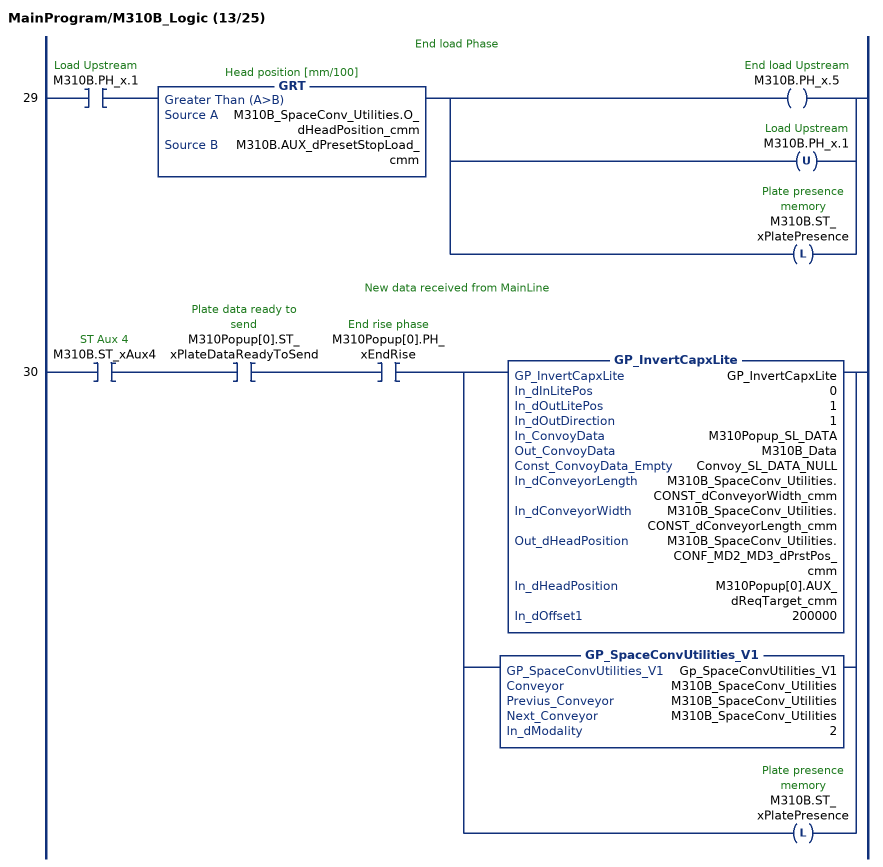
   // End load Phase
   29: XIC(M310B.PH_x.1)GRT(M310B_SpaceConv_Utilities.O_dHeadPosition_cmm,M310B.AUX_dPresetStopLoad_cmm)[OTE(M310B.PH_x.5) ,OTU(M310B.PH_x.1) ,OTL(M310B.ST_xPlatePresence) ];
   // New data received from MainLine
   30: XIC(M310B.ST_xAux4)XIC(M310Popup[0].ST_xPlateDataReadyToSend)XIC(M310Popup[0].PH_xEndRise)[GP_InvertCapxLite(GP_InvertCapxLite,0,1,1,M310Popup_SL_DATA,M310B_Data,Convoy_SL_DATA_NULL,M310B_SpaceConv_Utilities.CONST_dConveyorWidth_cmm,M310B_SpaceConv_Utilities.CONST_dConveyorLength_cmm,M310B_SpaceConv_Utilities.CONF_MD2_MD3_dPrstPos_cmm,M310Popup[0].AUX_dReqTarget_cmm,200000) ,GP_SpaceConvUtilities_V1(Gp_SpaceConvUtilities_V1,M310B_SpaceConv_Utilities,M310B_SpaceConv_Utilities,M310B_SpaceConv_Utilities,2) ,OTL(M310B.ST_xPlatePresence) ];
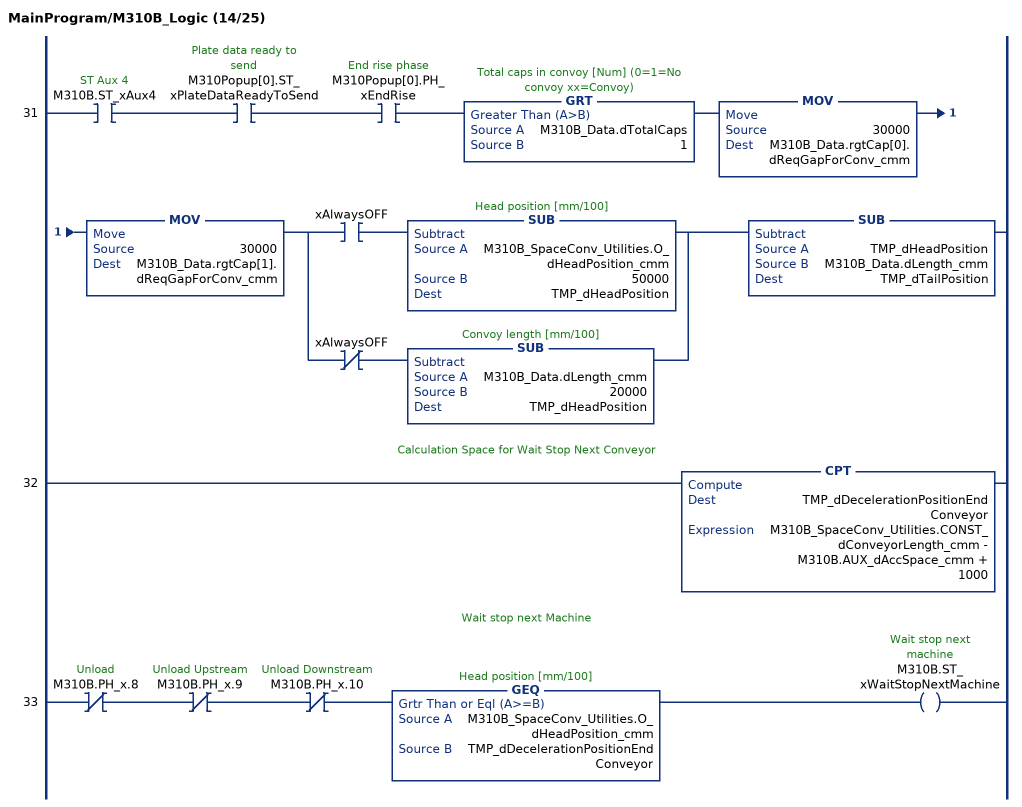
   31: XIC(M310B.ST_xAux4)XIC(M310Popup[0].ST_xPlateDataReadyToSend)XIC(M310Popup[0].PH_xEndRise)GRT(M310B_Data.dTotalCaps,1)MOV(30000,M310B_Data.rgtCap[0].dReqGapForConv_cmm)MOV(30000,M310B_Data.rgtCap[1].dReqGapForConv_cmm)[XIC(xAlwaysOFF) SUB(M310B_SpaceConv_Utilities.O_dHeadPosition_cmm,50000,TMP_dHeadPosition) ,XIO(xAlwaysOFF) SUB(M310B_Data.dLength_cmm,20000,TMP_dHeadPosition) ]SUB(TMP_dHeadPosition,M310B_Data.dLength_cmm,TMP_dTailPosition);
   // Calculation Space for Wait Stop Next Conveyor
   32: CPT(TMP_dDecelerationPositionEndConveyor,M310B_SpaceConv_Utilities.CONST_dConveyorLength_cmm - M310B.AUX_dAccSpace_cmm + 1000);
   // Wait stop next Machine
   33: XIO(M310B.PH_x.8)XIO(M310B.PH_x.9)XIO(M310B.PH_x.10)GEQ(M310B_SpaceConv_Utilities.O_dHeadPosition_cmm,TMP_dDecelerationPositionEndConveyor)OTE(M310B.ST_xWaitStopNextMachine);
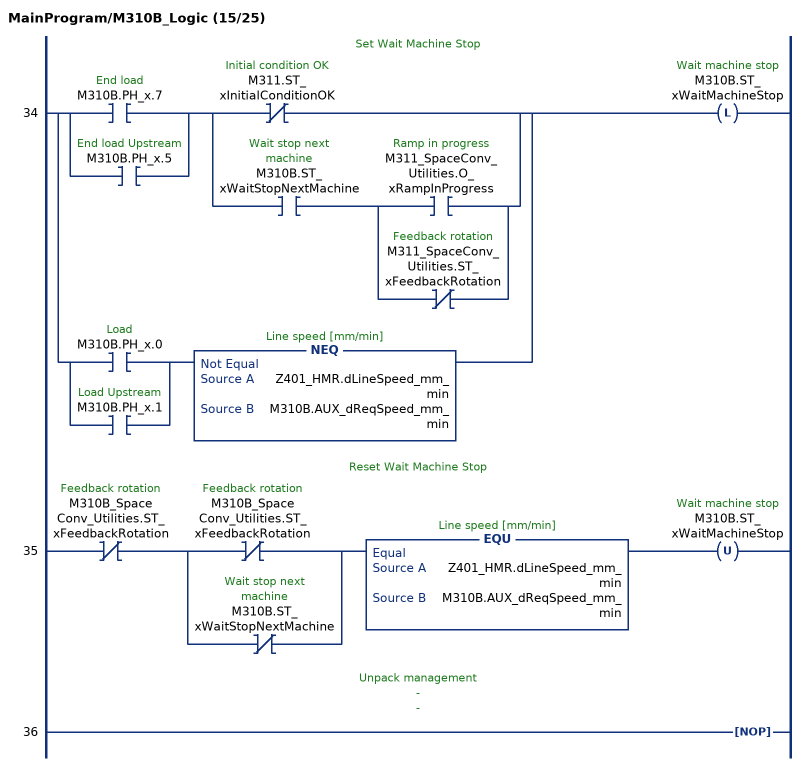
   // Set Wait Machine Stop
   34: [[XIC(M310B.PH_x.7) ,XIC(M310B.PH_x.5) ] [XIO(M311.ST_xInitialConditionOK) ,XIC(M310B.ST_xWaitStopNextMachine) [XIC(M311_SpaceConv_Utilities.O_xRampInProgress) ,XIO(M311_SpaceConv_Utilities.ST_xFeedbackRotation) ] ] ,[XIC(M310B.PH_x.0) ,XIC(M310B.PH_x.1) ] NEQ(Z401_HMR.dLineSpeed_mm_min,M310B.AUX_dReqSpeed_mm_min) ]OTL(M310B.ST_xWaitMachineStop);
   // Reset Wait Machine Stop
   35: XIO(M310B_SpaceConv_Utilities.ST_xFeedbackRotation)[XIO(M310B_SpaceConv_Utilities.ST_xFeedbackRotation) ,XIO(M310B.ST_xWaitStopNextMachine) ]EQU(Z401_HMR.dLineSpeed_mm_min,M310B.AUX_dReqSpeed_mm_min)OTU(M310B.ST_xWaitMachineStop);
   // Unpack management
   // -
   // -
   36: NOP();
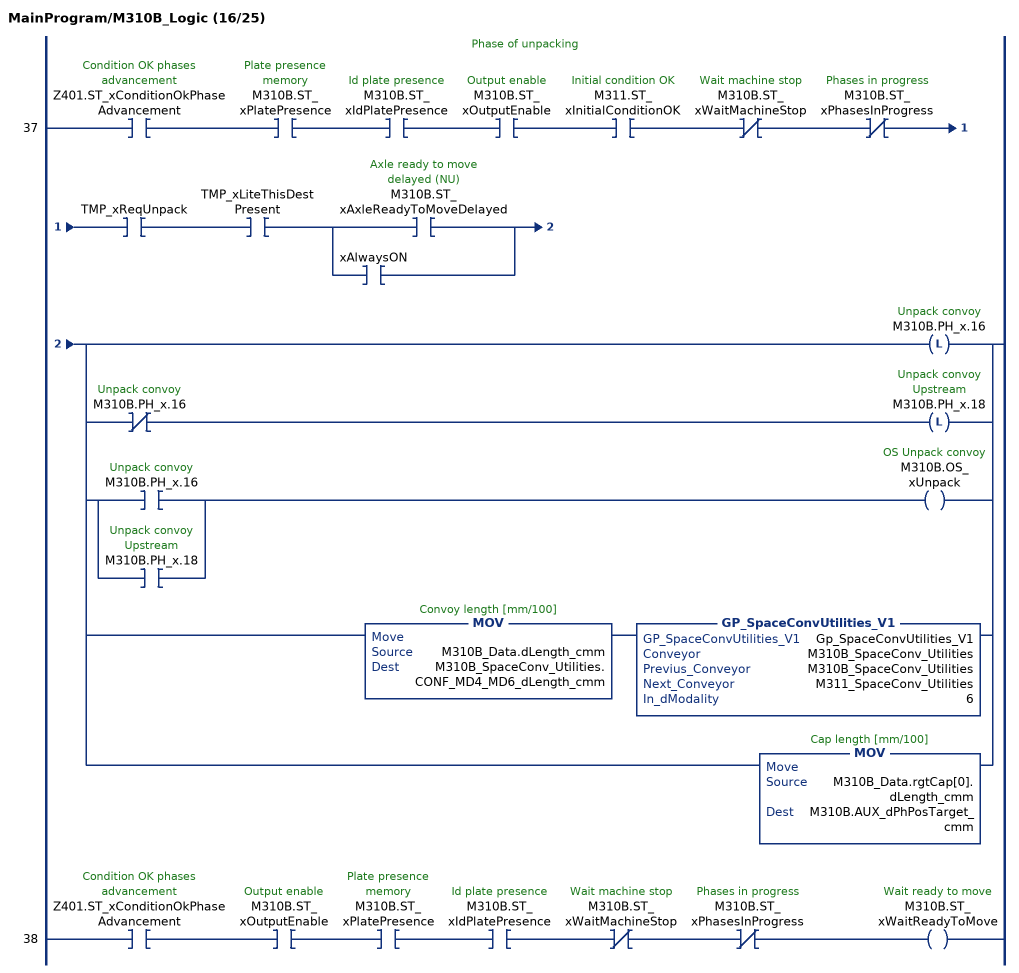
   // Phase of unpacking
   37: XIC(Z401.ST_xConditionOkPhaseAdvancement)XIC(M310B.ST_xPlatePresence)XIC(M310B.ST_xIdPlatePresence)XIC(M310B.ST_xOutputEnable)XIC(M311.ST_xInitialConditionOK)XIO(M310B.ST_xWaitMachineStop)XIO(M310B.ST_xPhasesInProgress)XIC(TMP_xReqUnpack)XIC(TMP_xLiteThisDestPresent)[XIC(M310B.ST_xAxleReadyToMoveDelayed) ,XIC(xAlwaysON) ][OTL(M310B.PH_x.16) ,XIO(M310B.PH_x.16) OTL(M310B.PH_x.18) ,[XIC(M310B.PH_x.16) ,XIC(M310B.PH_x.18) ] OTE(M310B.OS_xUnpack) ,MOV(M310B_Data.dLength_cmm,M310B_SpaceConv_Utilities.CONF_MD4_MD6_dLength_cmm) GP_SpaceConvUtilities_V1(Gp_SpaceConvUtilities_V1,M310B_SpaceConv_Utilities,M310B_SpaceConv_Utilities,M311_SpaceConv_Utilities,6) ,MOV(M310B_Data.rgtCap[0].dLength_cmm,M310B.AUX_dPhPosTarget_cmm) ];
   38: XIC(Z401.ST_xConditionOkPhaseAdvancement)XIC(M310B.ST_xOutputEnable)XIC(M310B.ST_xPlatePresence)XIC(M310B.ST_xIdPlatePresence)XIO(M310B.ST_xWaitMachineStop)XIO(M310B.ST_xPhasesInProgress)OTE(M310B.ST_xWaitReadyToMove);
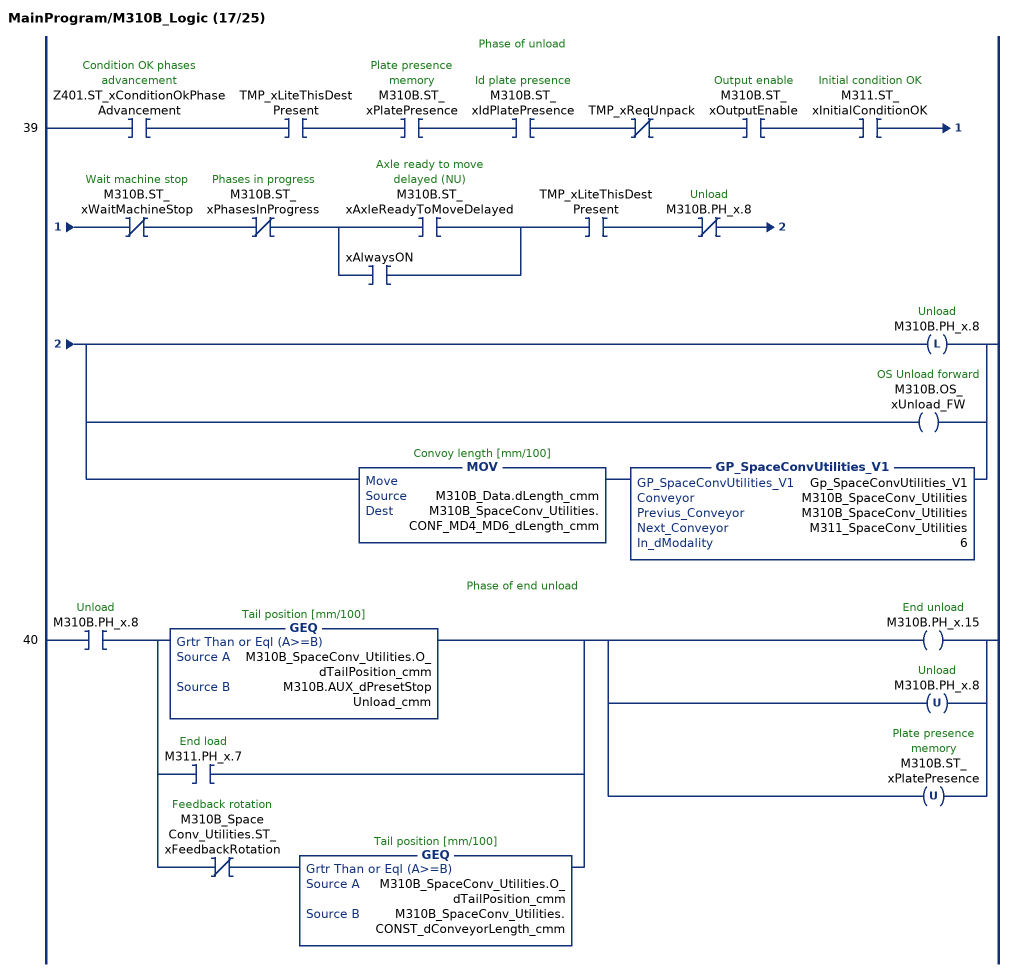
   // Phase of unload
   39: XIC(Z401.ST_xConditionOkPhaseAdvancement)XIC(TMP_xLiteThisDestPresent)XIC(M310B.ST_xPlatePresence)XIC(M310B.ST_xIdPlatePresence)XIO(TMP_xReqUnpack)XIC(M310B.ST_xOutputEnable)XIC(M311.ST_xInitialConditionOK)XIO(M310B.ST_xWaitMachineStop)XIO(M310B.ST_xPhasesInProgress)[XIC(M310B.ST_xAxleReadyToMoveDelayed) ,XIC(xAlwaysON) ]XIC(TMP_xLiteThisDestPresent)XIO(M310B.PH_x.8)[OTL(M310B.PH_x.8) ,OTE(M310B.OS_xUnload_FW) ,MOV(M310B_Data.dLength_cmm,M310B_SpaceConv_Utilities.CONF_MD4_MD6_dLength_cmm) GP_SpaceConvUtilities_V1(Gp_SpaceConvUtilities_V1,M310B_SpaceConv_Utilities,M310B_SpaceConv_Utilities,M311_SpaceConv_Utilities,6) ];
   // Phase of end unload
   40: XIC(M310B.PH_x.8)[[GEQ(M310B_SpaceConv_Utilities.O_dTailPosition_cmm,M310B.AUX_dPresetStopUnload_cmm) ,XIC(M311.PH_x.7) ] ,XIO(M310B_SpaceConv_Utilities.ST_xFeedbackRotation) GEQ(M310B_SpaceConv_Utilities.O_dTailPosition_cmm,M310B_SpaceConv_Utilities.CONST_dConveyorLength_cmm) ][OTE(M310B.PH_x.15) ,OTU(M310B.PH_x.8) ,OTU(M310B.ST_xPlatePresence) ];
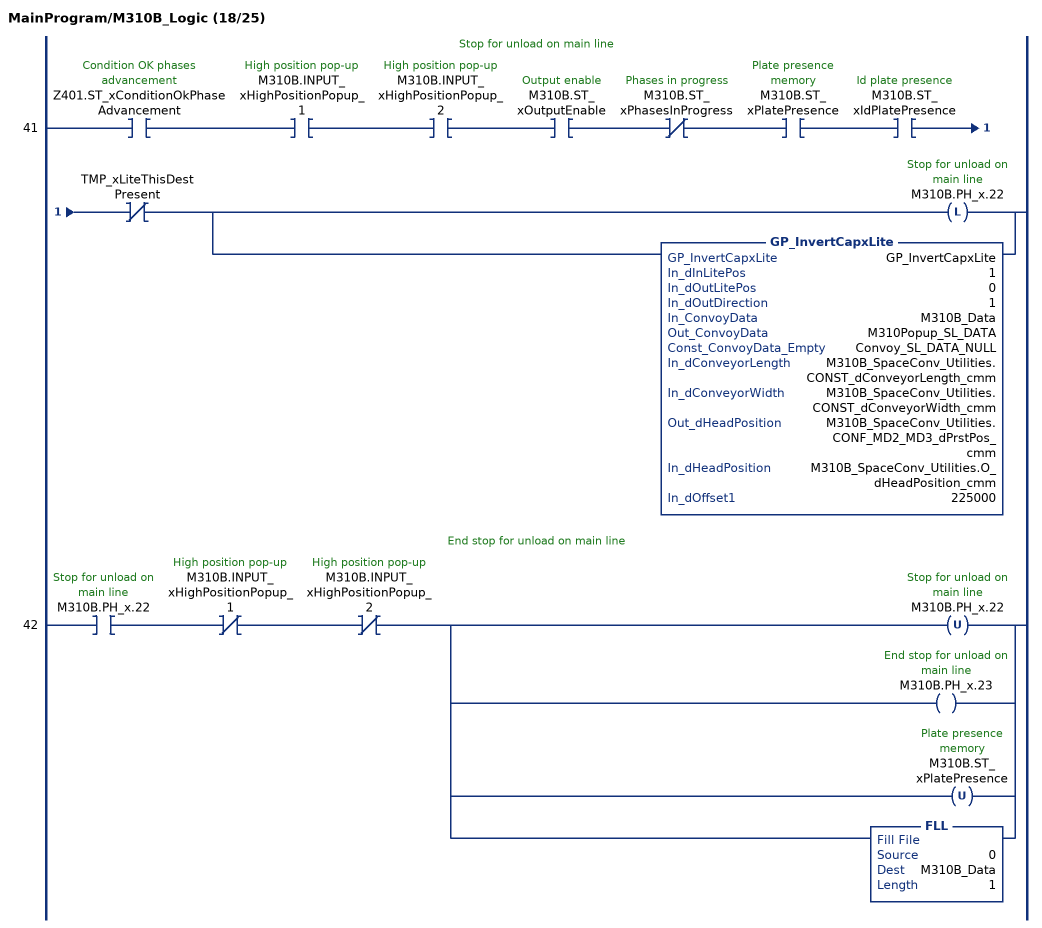
   // Stop for unload on main line
   41: XIC(Z401.ST_xConditionOkPhaseAdvancement)XIC(M310B.INPUT_xHighPositionPopup_1)XIC(M310B.INPUT_xHighPositionPopup_2)XIC(M310B.ST_xOutputEnable)XIO(M310B.ST_xPhasesInProgress)XIC(M310B.ST_xPlatePresence)XIC(M310B.ST_xIdPlatePresence)XIO(TMP_xLiteThisDestPresent)[OTL(M310B.PH_x.22) ,GP_InvertCapxLite(GP_InvertCapxLite,1,0,1,M310B_Data,M310Popup_SL_DATA,Convoy_SL_DATA_NULL,M310B_SpaceConv_Utilities.CONST_dConveyorLength_cmm,M310B_SpaceConv_Utilities.CONST_dConveyorWidth_cmm,M310B_SpaceConv_Utilities.CONF_MD2_MD3_dPrstPos_cmm,M310B_SpaceConv_Utilities.O_dHeadPosition_cmm,225000) ];
   // End stop for unload on main line
   42: XIC(M310B.PH_x.22)XIO(M310B.INPUT_xHighPositionPopup_1)XIO(M310B.INPUT_xHighPositionPopup_2)[OTU(M310B.PH_x.22) ,OTE(M310B.PH_x.23) ,OTU(M310B.ST_xPlatePresence) ,FLL(0,M310B_Data,1) ];
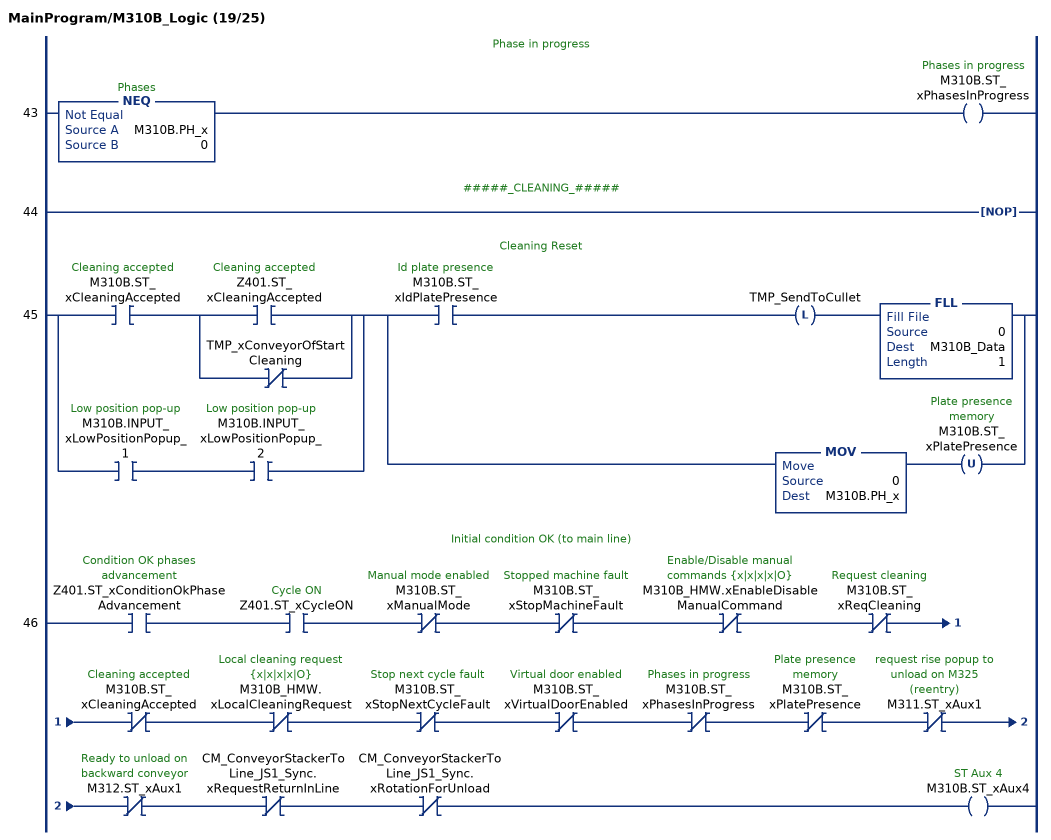
   // Phase in progress
   43: NEQ(M310B.PH_x,0)OTE(M310B.ST_xPhasesInProgress);
   // #####_CLEANING_#####
   44: NOP();
   // Cleaning Reset
   45: [XIC(M310B.ST_xCleaningAccepted) [XIC(Z401.ST_xCleaningAccepted) ,XIO(TMP_xConveyorOfStartCleaning) ] ,XIC(M310B.INPUT_xLowPositionPopup_1) XIC(M310B.INPUT_xLowPositionPopup_2) ][XIC(M310B.ST_xIdPlatePresence) OTL(TMP_SendToCullet) FLL(0,M310B_Data,1) ,MOV(0,M310B.PH_x) OTU(M310B.ST_xPlatePresence) ];
   // Initial condition OK (to main line)
   46: XIC(Z401.ST_xConditionOkPhaseAdvancement)XIC(Z401.ST_xCycleON)XIO(M310B.ST_xManualMode)XIO(M310B.ST_xStopMachineFault)XIO(M310B_HMW.xEnableDisableManualCommand)XIO(M310B.ST_xReqCleaning)XIO(M310B.ST_xCleaningAccepted)XIO(M310B_HMW.xLocalCleaningRequest)XIO(M310B.ST_xStopNextCycleFault)XIO(M310B.ST_xVirtualDoorEnabled)XIO(M310B.ST_xPhasesInProgress)XIO(M310B.ST_xPlatePresence)XIO(M311.ST_xAux1)XIO(M312.ST_xAux1)XIO(CM_ConveyorStackerToLine_JS1_Sync.xRequestReturnInLine)XIO(CM_ConveyorStackerToLine_JS1_Sync.xRotationForUnload)OTE(M310B.ST_xAux4);
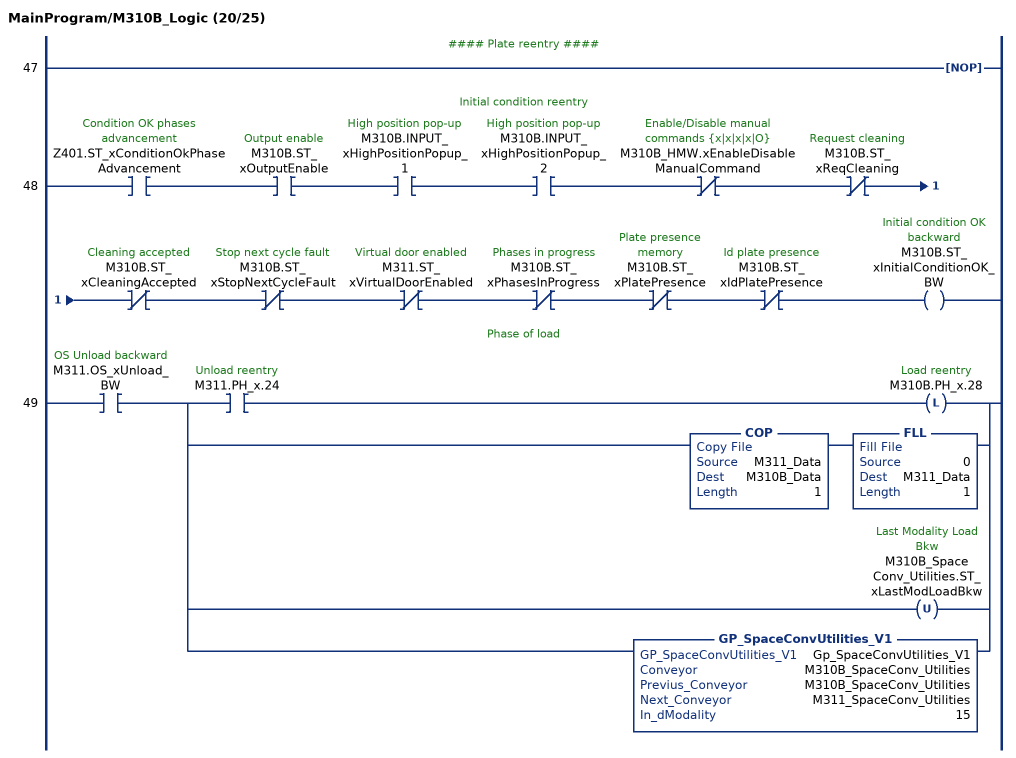
   // #### Plate reentry ####
   47: NOP();
   // Initial condition reentry
   48: XIC(Z401.ST_xConditionOkPhaseAdvancement)XIC(M310B.ST_xOutputEnable)XIC(M310B.INPUT_xHighPositionPopup_1)XIC(M310B.INPUT_xHighPositionPopup_2)XIO(M310B_HMW.xEnableDisableManualCommand)XIO(M310B.ST_xReqCleaning)XIO(M310B.ST_xCleaningAccepted)XIO(M310B.ST_xStopNextCycleFault)XIO(M311.ST_xVirtualDoorEnabled)XIO(M310B.ST_xPhasesInProgress)XIO(M310B.ST_xPlatePresence)XIO(M310B.ST_xIdPlatePresence)OTE(M310B.ST_xInitialConditionOK_BW);
   // Phase of load
   49: XIC(M311.OS_xUnload_BW)[XIC(M311.PH_x.24) OTL(M310B.PH_x.28) ,COP(M311_Data,M310B_Data,1) FLL(0,M311_Data,1) ,OTU(M310B_SpaceConv_Utilities.ST_xLastModLoadBkw) ,GP_SpaceConvUtilities_V1(Gp_SpaceConvUtilities_V1,M310B_SpaceConv_Utilities,M310B_SpaceConv_Utilities,M311_SpaceConv_Utilities,15) ];
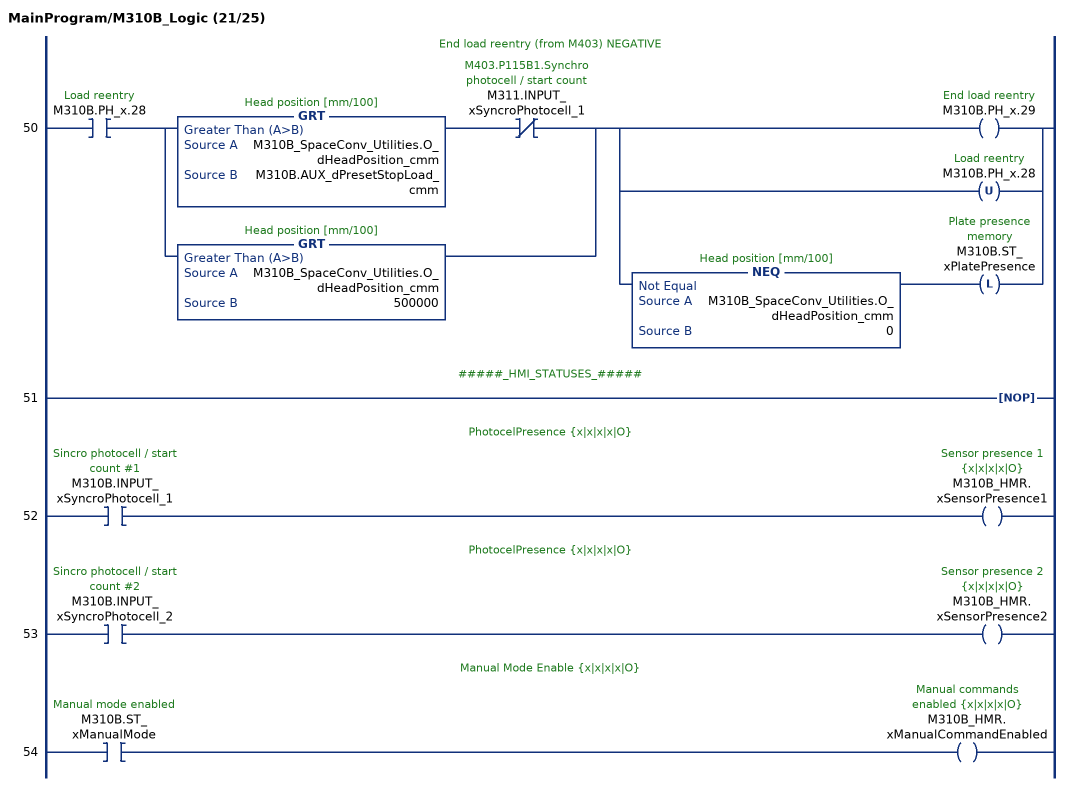
   // End load reentry (from M403) NEGATIVE
   50: XIC(M310B.PH_x.28)[GRT(M310B_SpaceConv_Utilities.O_dHeadPosition_cmm,M310B.AUX_dPresetStopLoad_cmm) XIO(M311.INPUT_xSyncroPhotocell_1) ,GRT(M310B_SpaceConv_Utilities.O_dHeadPosition_cmm,500000) ][OTE(M310B.PH_x.29) ,OTU(M310B.PH_x.28) ,NEQ(M310B_SpaceConv_Utilities.O_dHeadPosition_cmm,0) OTL(M310B.ST_xPlatePresence) ];
   // #####_HMI_STATUSES_#####
   51: NOP();
   // PhotocelPresence {x|x|x|x|O}
   52: XIC(M310B.INPUT_xSyncroPhotocell_1)OTE(M310B_HMR.xSensorPresence1);
   // PhotocelPresence {x|x|x|x|O}
   53: XIC(M310B.INPUT_xSyncroPhotocell_2)OTE(M310B_HMR.xSensorPresence2);
   // Manual Mode Enable {x|x|x|x|O}
   54: XIC(M310B.ST_xManualMode)OTE(M310B_HMR.xManualCommandEnabled);
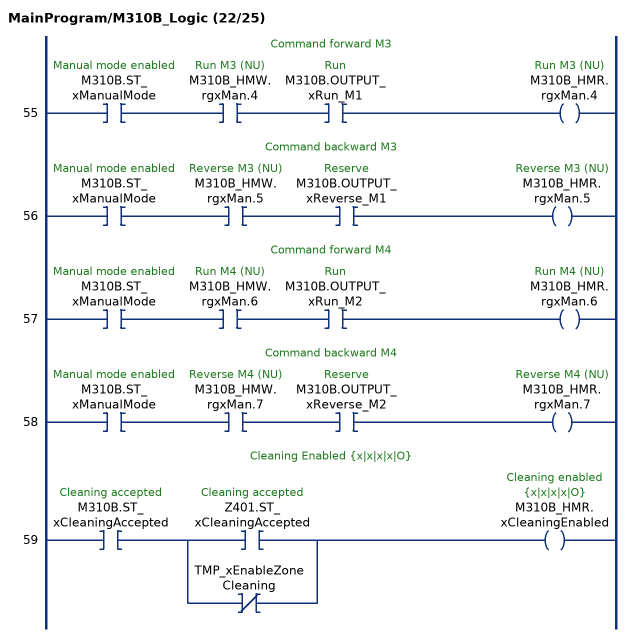
   // Command forward M3
   55: XIC(M310B.ST_xManualMode)XIC(M310B_HMW.rgxMan.4)XIC(M310B.OUTPUT_xRun_M1)OTE(M310B_HMR.rgxMan.4);
   // Command backward M3
   56: XIC(M310B.ST_xManualMode)XIC(M310B_HMW.rgxMan.5)XIC(M310B.OUTPUT_xReverse_M1)OTE(M310B_HMR.rgxMan.5);
   // Command forward M4
   57: XIC(M310B.ST_xManualMode)XIC(M310B_HMW.rgxMan.6)XIC(M310B.OUTPUT_xRun_M2)OTE(M310B_HMR.rgxMan.6);
   // Command backward M4
   58: XIC(M310B.ST_xManualMode)XIC(M310B_HMW.rgxMan.7)XIC(M310B.OUTPUT_xReverse_M2)OTE(M310B_HMR.rgxMan.7);
   // Cleaning Enabled {x|x|x|x|O}
   59: XIC(M310B.ST_xCleaningAccepted)[XIC(Z401.ST_xCleaningAccepted) ,XIO(TMP_xEnableZoneCleaning) ]OTE(M310B_HMR.xCleaningEnabled);
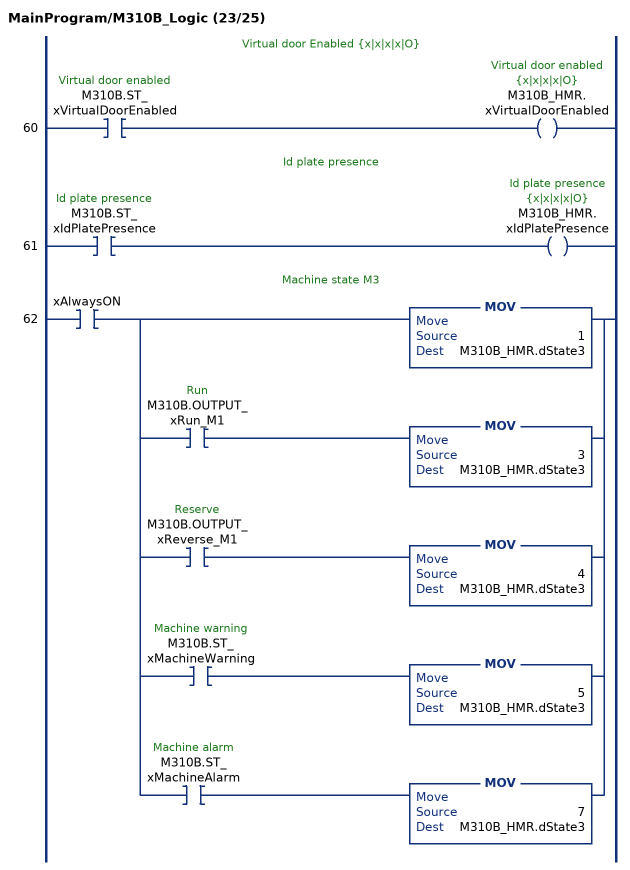
   // Virtual door Enabled {x|x|x|x|O}
   60: XIC(M310B.ST_xVirtualDoorEnabled)OTE(M310B_HMR.xVirtualDoorEnabled);
   // Id plate presence
   61: XIC(M310B.ST_xIdPlatePresence)OTE(M310B_HMR.xIdPlatePresence);
   // Machine state M3
   62: XIC(xAlwaysON)[MOV(1,M310B_HMR.dState3) ,XIC(M310B.OUTPUT_xRun_M1) MOV(3,M310B_HMR.dState3) ,XIC(M310B.OUTPUT_xReverse_M1) MOV(4,M310B_HMR.dState3) ,XIC(M310B.ST_xMachineWarning) MOV(5,M310B_HMR.dState3) ,XIC(M310B.ST_xMachineAlarm) MOV(7,M310B_HMR.dState3) ];
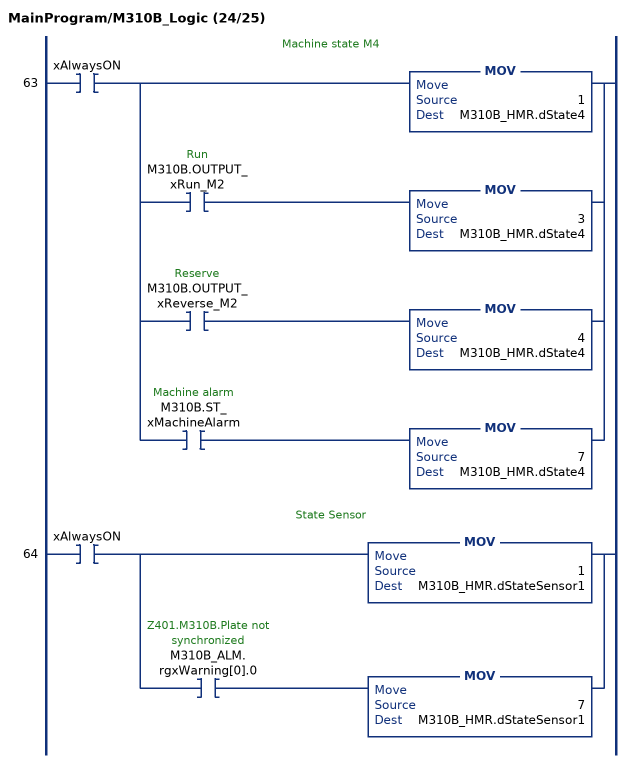
   // Machine state M4
   63: XIC(xAlwaysON)[MOV(1,M310B_HMR.dState4) ,XIC(M310B.OUTPUT_xRun_M2) MOV(3,M310B_HMR.dState4) ,XIC(M310B.OUTPUT_xReverse_M2) MOV(4,M310B_HMR.dState4) ,XIC(M310B.ST_xMachineAlarm) MOV(7,M310B_HMR.dState4) ];
   // State Sensor
   64: XIC(xAlwaysON)[MOV(1,M310B_HMR.dStateSensor1) ,XIC(M310B_ALM.rgxWarning[0].0) MOV(7,M310B_HMR.dStateSensor1) ];
